(* Logix 5000 project; controller MV vendor 1 type 14 code 217 rev 31.11; software revision 31.00; part 50 of 53 *)
(* tags used below, declared in another part *)
   CC_CIP_BeerMain_Active : DINT;
   CheckTimeMask : INT;
   Delphi_Does_Eng_Func : BOOL;
   enable_comms_to_fv_plc : BOOL;
   MV_BM01_AV01_CIP : BOOL;
   mv_comms_from_cc_plc : MESSAGE;
   mv_comms_from_cc_timer : TIMER;
   MV_COMMS_FROM_FV_PLC : MESSAGE;
   mv_comms_from_mv_routing_plc : MESSAGE;
   mv_comms_to_fv_plc : MESSAGE;
   mv_comms_to_fv_plc_timer : TIMER;
   mv_comms_to_mv_routing_plc : MESSAGE;
   mv_comms_to_mv_routing_plc_timer : TIMER;
   MV_data_file_value_to_move : DINT;
   MV_MV10R : PlantItem;   // MV10R
   MV_MV11R : PlantItem;   // MV11R
   MV_MV12R : PlantItem;   // MV12R
   MV_MV13R : PlantItem;   // MV13R
   MV_MV14R : PlantItem;   // MV14R
   MV_MV15R : PlantItem;   // MV15R
   MV_MV16R : PlantItem;   // MV16R
   MV_MV17R : PlantItem;   // MV17R
   MV_MV18R : PlantItem;   // MV18R
   MV_MV19R : PlantItem;   // MV19R
   MV_MV20_TP_KBEmptying : BOOL;
   MV_MV20R : PlantItem;   // MV20R
   MV_MV21_TP_KBEmptying : BOOL;
   MV_MV21R : PlantItem;   // MV21R
   MV_MV22_TP_KBEmptying : BOOL;
   MV_MV22R : PlantItem;   // MV22R
   MV_MV23R : PlantItem;   // MV23R
   MV_MV30R : PlantItem;   // MV30R
   MV_MV31R : PlantItem;   // MV31R
   MV_MV32R : PlantItem;   // MV32R
   MV_MV33R : PlantItem;   // MV33R
   MV_MV34R : PlantItem;   // MV34R
   MV_MV35R : PlantItem;   // MV35R
   MV_MV7R : PlantItem;   // MV7R
   MV_MV8R : PlantItem;   // MV8R
   MV_MV9R : PlantItem;   // MV9R
   MV_N13 : INT[255];   // PLC>ME Inter PLC comms traf fic inbound
   MV_N14 : INT[255];   // ME>PLC Inter PLC comms traf fic outbound
   MV_N140 : INT[50];   // MV 36, CURRENT FV DATA
   MV_N141 : INT[50];   // MV 37, CURRENT FV DATA
   MV_N142 : INT[50];   // MV 38, CURRENT FV DATA
   MV_N143 : INT[50];   // MV 39, CURRENT FV DATA
   MV_N144 : INT[50];   // MV 40, CURRENT FV DATA
   MV_N145 : INT[50];   // MV 41, CURRENT FV DATA
   MV_N146 : INT[50];   // MV 42, CURRENT FV DATA
   MV_N147 : INT[50];   // MV 43, CURRENT FV DATA
   MV_N148 : INT[50];   // MV 44, CURRENT FV DATA
   MV_N149 : INT[50];   // MV 45, CURRENT FV DATA
   MV_N15 : INT[255];   // COMMS_CTRL Inter PLC comms inte rnal working regs
   MV_N150 : INT[50];   // MV 36, CURRENT FV DATA
   MV_N151 : INT[50];   // MV 47, CURRENT FV DATA
   MV_N15_63_0_OutputBit : BOOL;
   MV_N190 : INT[255];   // Original N File From SLC, No Description Available
   MV_N255 : DINT[255];   // Old Format Checkwords To Keep Delphi Indicating Status Correctly.
   MV_T16 : TIMER[10];
   MV_T191 : TIMER[20];
   MV_T4 : TIMER[20];
   TempChecktime : DINT;
(* MV_Common, continued *)

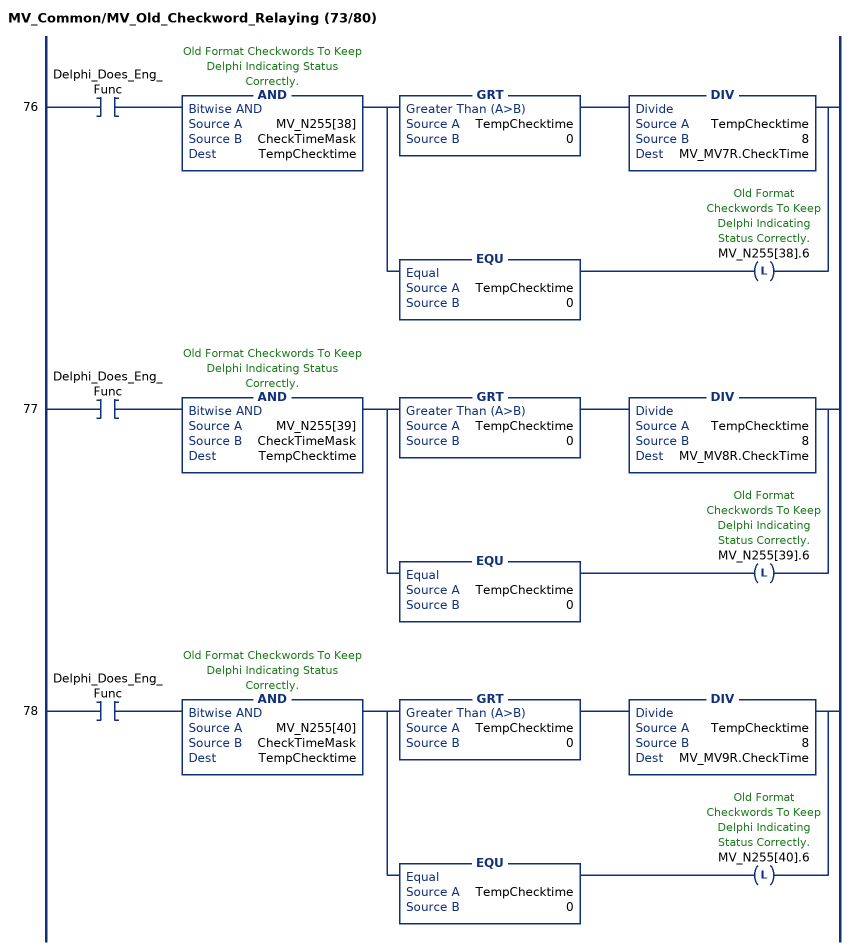
   [picture p1231: MV_Common/MV_Old_Checkword_Relaying rungs 76-78]
   76: XIC(Delphi_Does_Eng_Func)AND(MV_N255[38],CheckTimeMask,TempChecktime)[GRT(TempChecktime,0) DIV(TempChecktime,8,MV_MV7R.CheckTime) ,EQU(TempChecktime,0) OTL(MV_N255[38].6) ];
   77: XIC(Delphi_Does_Eng_Func)AND(MV_N255[39],CheckTimeMask,TempChecktime)[GRT(TempChecktime,0) DIV(TempChecktime,8,MV_MV8R.CheckTime) ,EQU(TempChecktime,0) OTL(MV_N255[39].6) ];
   78: XIC(Delphi_Does_Eng_Func)AND(MV_N255[40],CheckTimeMask,TempChecktime)[GRT(TempChecktime,0) DIV(TempChecktime,8,MV_MV9R.CheckTime) ,EQU(TempChecktime,0) OTL(MV_N255[40].6) ];
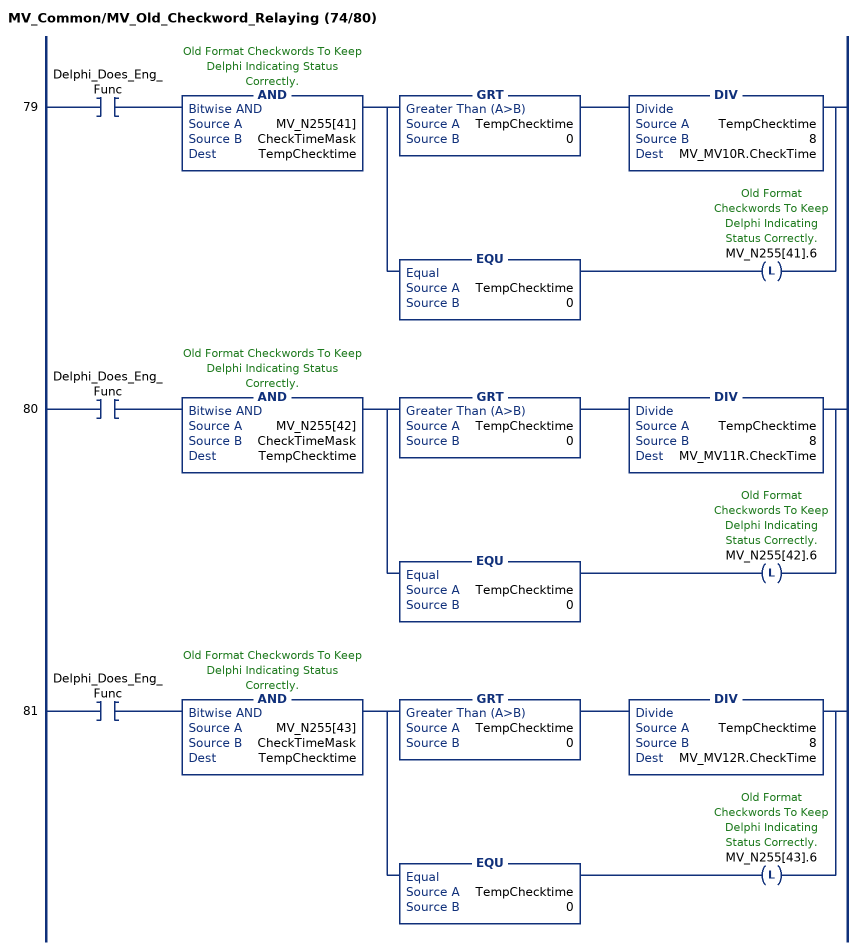
   79: XIC(Delphi_Does_Eng_Func)AND(MV_N255[41],CheckTimeMask,TempChecktime)[GRT(TempChecktime,0) DIV(TempChecktime,8,MV_MV10R.CheckTime) ,EQU(TempChecktime,0) OTL(MV_N255[41].6) ];
   80: XIC(Delphi_Does_Eng_Func)AND(MV_N255[42],CheckTimeMask,TempChecktime)[GRT(TempChecktime,0) DIV(TempChecktime,8,MV_MV11R.CheckTime) ,EQU(TempChecktime,0) OTL(MV_N255[42].6) ];
   81: XIC(Delphi_Does_Eng_Func)AND(MV_N255[43],CheckTimeMask,TempChecktime)[GRT(TempChecktime,0) DIV(TempChecktime,8,MV_MV12R.CheckTime) ,EQU(TempChecktime,0) OTL(MV_N255[43].6) ];
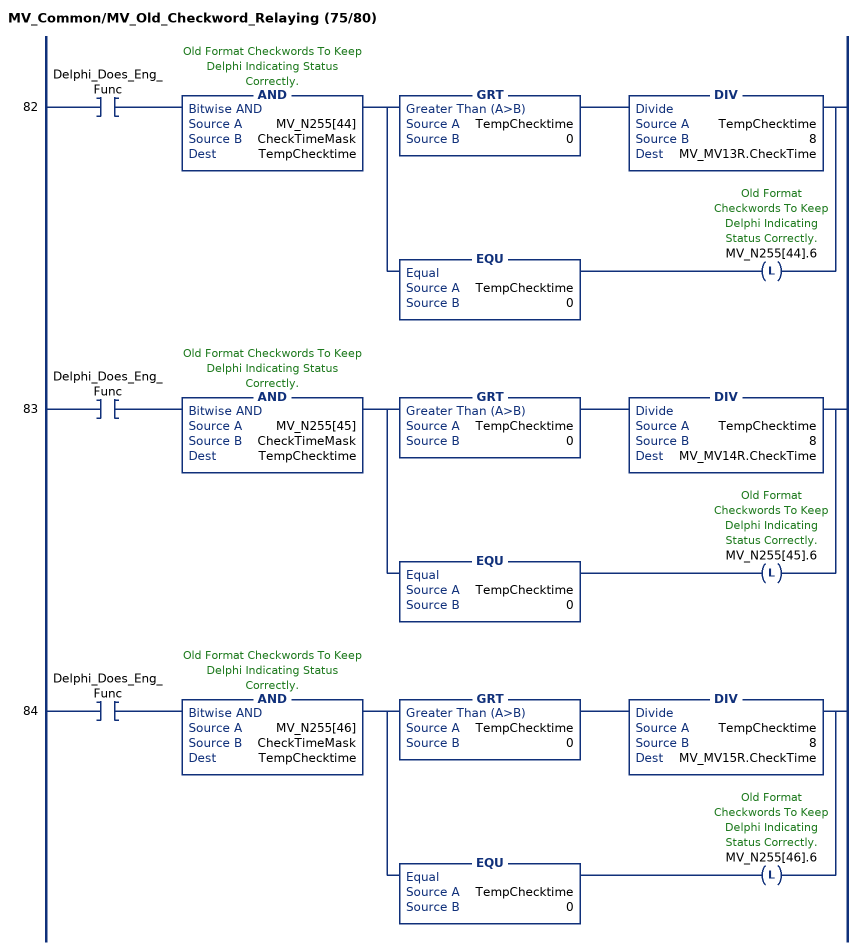
   82: XIC(Delphi_Does_Eng_Func)AND(MV_N255[44],CheckTimeMask,TempChecktime)[GRT(TempChecktime,0) DIV(TempChecktime,8,MV_MV13R.CheckTime) ,EQU(TempChecktime,0) OTL(MV_N255[44].6) ];
   83: XIC(Delphi_Does_Eng_Func)AND(MV_N255[45],CheckTimeMask,TempChecktime)[GRT(TempChecktime,0) DIV(TempChecktime,8,MV_MV14R.CheckTime) ,EQU(TempChecktime,0) OTL(MV_N255[45].6) ];
   84: XIC(Delphi_Does_Eng_Func)AND(MV_N255[46],CheckTimeMask,TempChecktime)[GRT(TempChecktime,0) DIV(TempChecktime,8,MV_MV15R.CheckTime) ,EQU(TempChecktime,0) OTL(MV_N255[46].6) ];
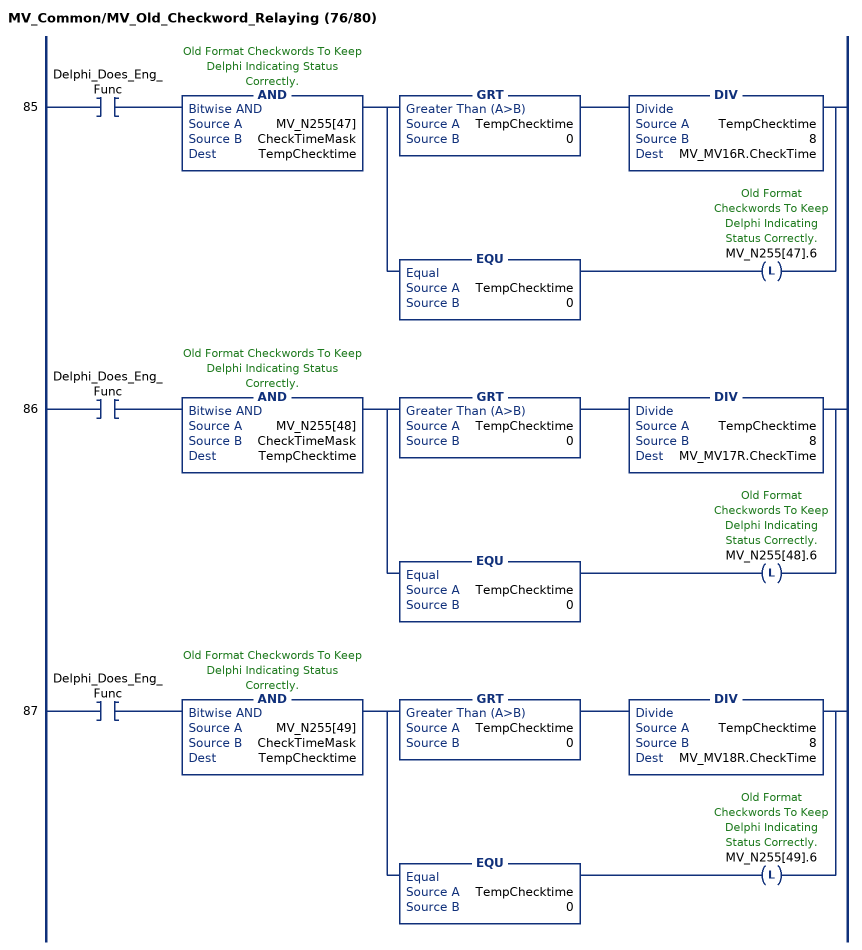
   85: XIC(Delphi_Does_Eng_Func)AND(MV_N255[47],CheckTimeMask,TempChecktime)[GRT(TempChecktime,0) DIV(TempChecktime,8,MV_MV16R.CheckTime) ,EQU(TempChecktime,0) OTL(MV_N255[47].6) ];
   86: XIC(Delphi_Does_Eng_Func)AND(MV_N255[48],CheckTimeMask,TempChecktime)[GRT(TempChecktime,0) DIV(TempChecktime,8,MV_MV17R.CheckTime) ,EQU(TempChecktime,0) OTL(MV_N255[48].6) ];
   87: XIC(Delphi_Does_Eng_Func)AND(MV_N255[49],CheckTimeMask,TempChecktime)[GRT(TempChecktime,0) DIV(TempChecktime,8,MV_MV18R.CheckTime) ,EQU(TempChecktime,0) OTL(MV_N255[49].6) ];
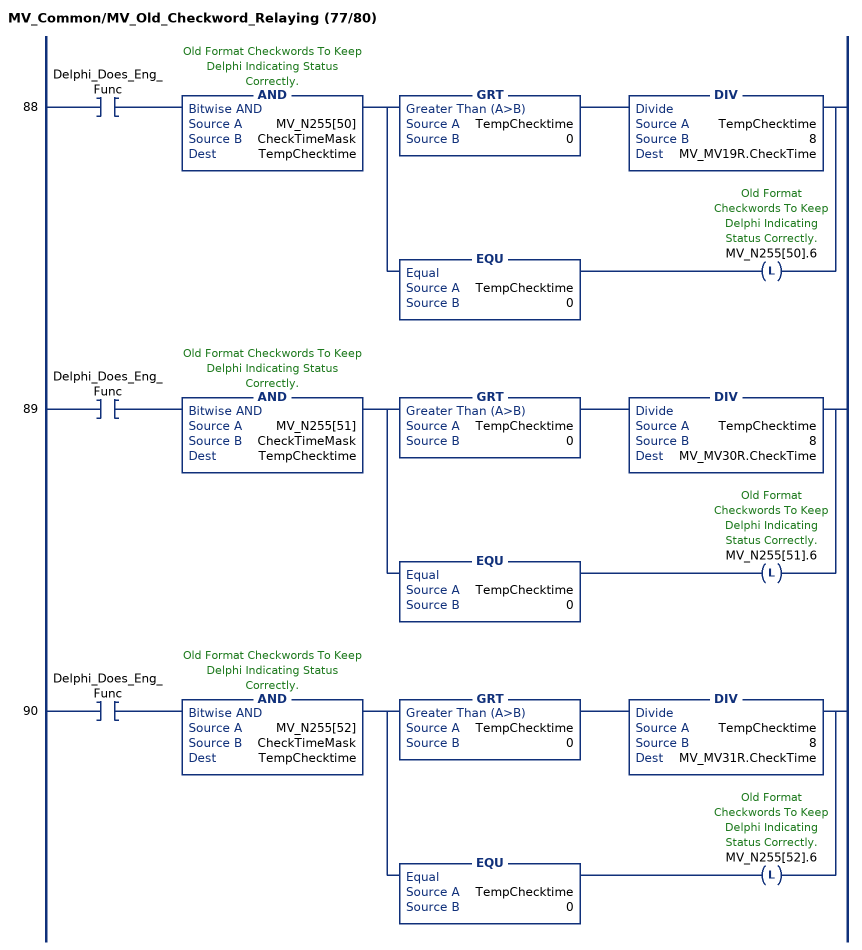
   88: XIC(Delphi_Does_Eng_Func)AND(MV_N255[50],CheckTimeMask,TempChecktime)[GRT(TempChecktime,0) DIV(TempChecktime,8,MV_MV19R.CheckTime) ,EQU(TempChecktime,0) OTL(MV_N255[50].6) ];
   89: XIC(Delphi_Does_Eng_Func)AND(MV_N255[51],CheckTimeMask,TempChecktime)[GRT(TempChecktime,0) DIV(TempChecktime,8,MV_MV30R.CheckTime) ,EQU(TempChecktime,0) OTL(MV_N255[51].6) ];
   90: XIC(Delphi_Does_Eng_Func)AND(MV_N255[52],CheckTimeMask,TempChecktime)[GRT(TempChecktime,0) DIV(TempChecktime,8,MV_MV31R.CheckTime) ,EQU(TempChecktime,0) OTL(MV_N255[52].6) ];
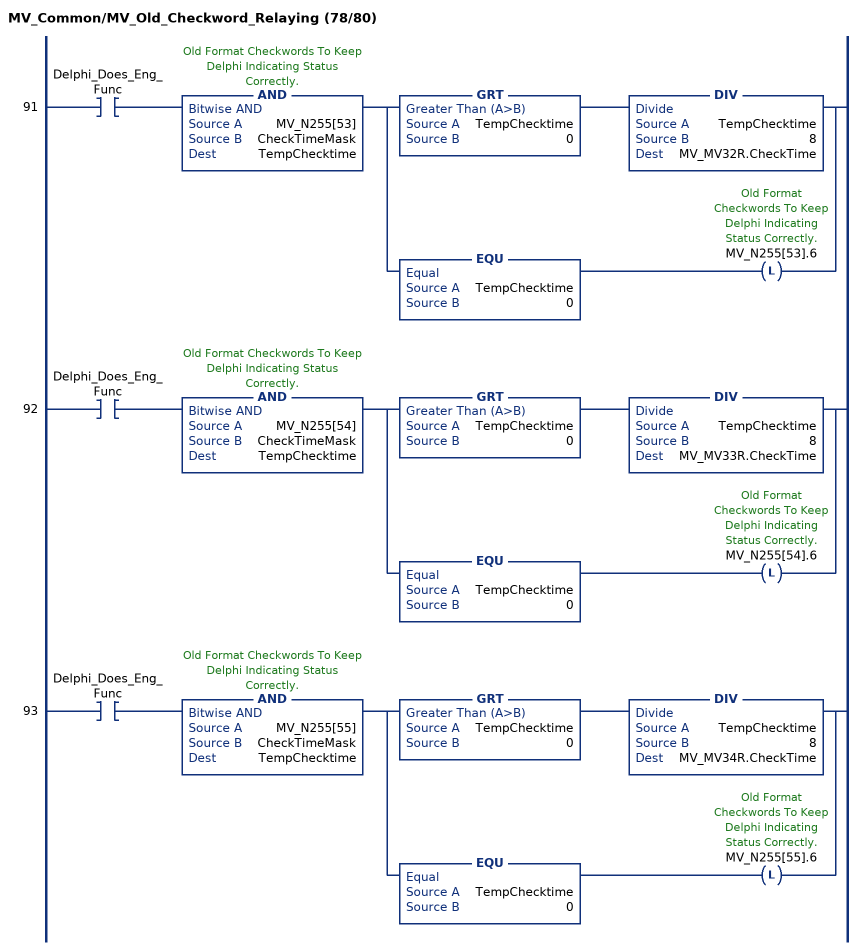
   91: XIC(Delphi_Does_Eng_Func)AND(MV_N255[53],CheckTimeMask,TempChecktime)[GRT(TempChecktime,0) DIV(TempChecktime,8,MV_MV32R.CheckTime) ,EQU(TempChecktime,0) OTL(MV_N255[53].6) ];
   92: XIC(Delphi_Does_Eng_Func)AND(MV_N255[54],CheckTimeMask,TempChecktime)[GRT(TempChecktime,0) DIV(TempChecktime,8,MV_MV33R.CheckTime) ,EQU(TempChecktime,0) OTL(MV_N255[54].6) ];
   93: XIC(Delphi_Does_Eng_Func)AND(MV_N255[55],CheckTimeMask,TempChecktime)[GRT(TempChecktime,0) DIV(TempChecktime,8,MV_MV34R.CheckTime) ,EQU(TempChecktime,0) OTL(MV_N255[55].6) ];
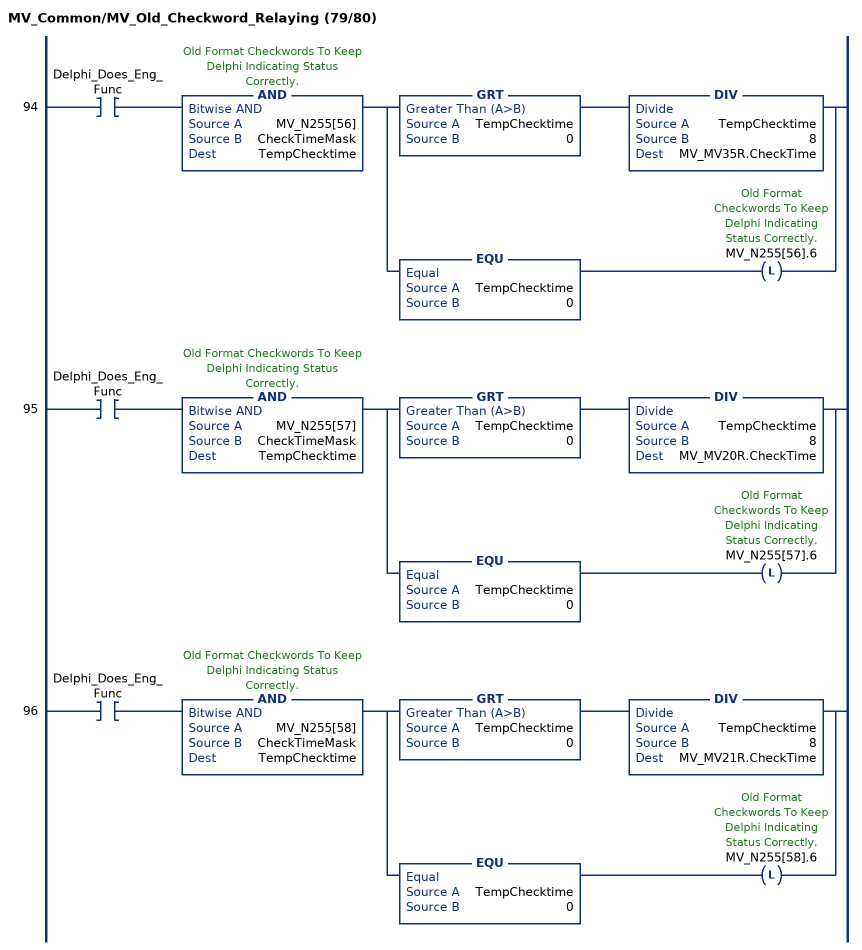
   94: XIC(Delphi_Does_Eng_Func)AND(MV_N255[56],CheckTimeMask,TempChecktime)[GRT(TempChecktime,0) DIV(TempChecktime,8,MV_MV35R.CheckTime) ,EQU(TempChecktime,0) OTL(MV_N255[56].6) ];
   95: XIC(Delphi_Does_Eng_Func)AND(MV_N255[57],CheckTimeMask,TempChecktime)[GRT(TempChecktime,0) DIV(TempChecktime,8,MV_MV20R.CheckTime) ,EQU(TempChecktime,0) OTL(MV_N255[57].6) ];
   96: XIC(Delphi_Does_Eng_Func)AND(MV_N255[58],CheckTimeMask,TempChecktime)[GRT(TempChecktime,0) DIV(TempChecktime,8,MV_MV21R.CheckTime) ,EQU(TempChecktime,0) OTL(MV_N255[58].6) ];
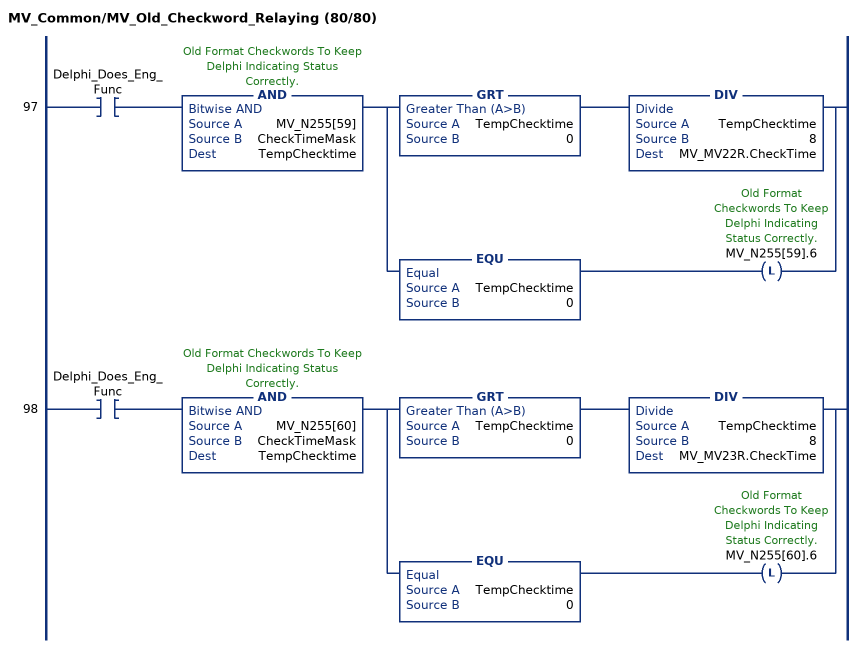
   97: XIC(Delphi_Does_Eng_Func)AND(MV_N255[59],CheckTimeMask,TempChecktime)[GRT(TempChecktime,0) DIV(TempChecktime,8,MV_MV22R.CheckTime) ,EQU(TempChecktime,0) OTL(MV_N255[59].6) ];
   98: XIC(Delphi_Does_Eng_Func)AND(MV_N255[60],CheckTimeMask,TempChecktime)[GRT(TempChecktime,0) DIV(TempChecktime,8,MV_MV23R.CheckTime) ,EQU(TempChecktime,0) OTL(MV_N255[60].6) ];
END_ROUTINE

ROUTINE MV_PLC_COMMS_7   (* ladder *)
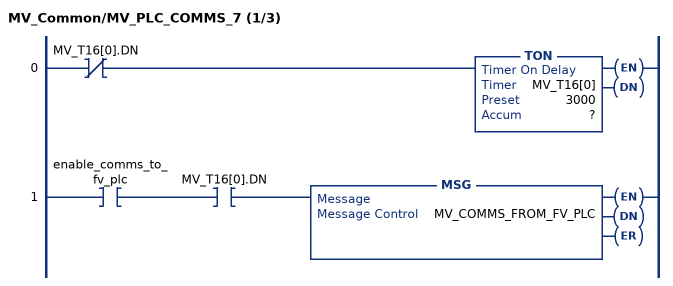
   0: XIO(MV_T16[0].DN)TON(MV_T16[0],?,?);
   1: XIC(enable_comms_to_fv_plc)XIC(MV_T16[0].DN)MSG(MV_COMMS_FROM_FV_PLC);
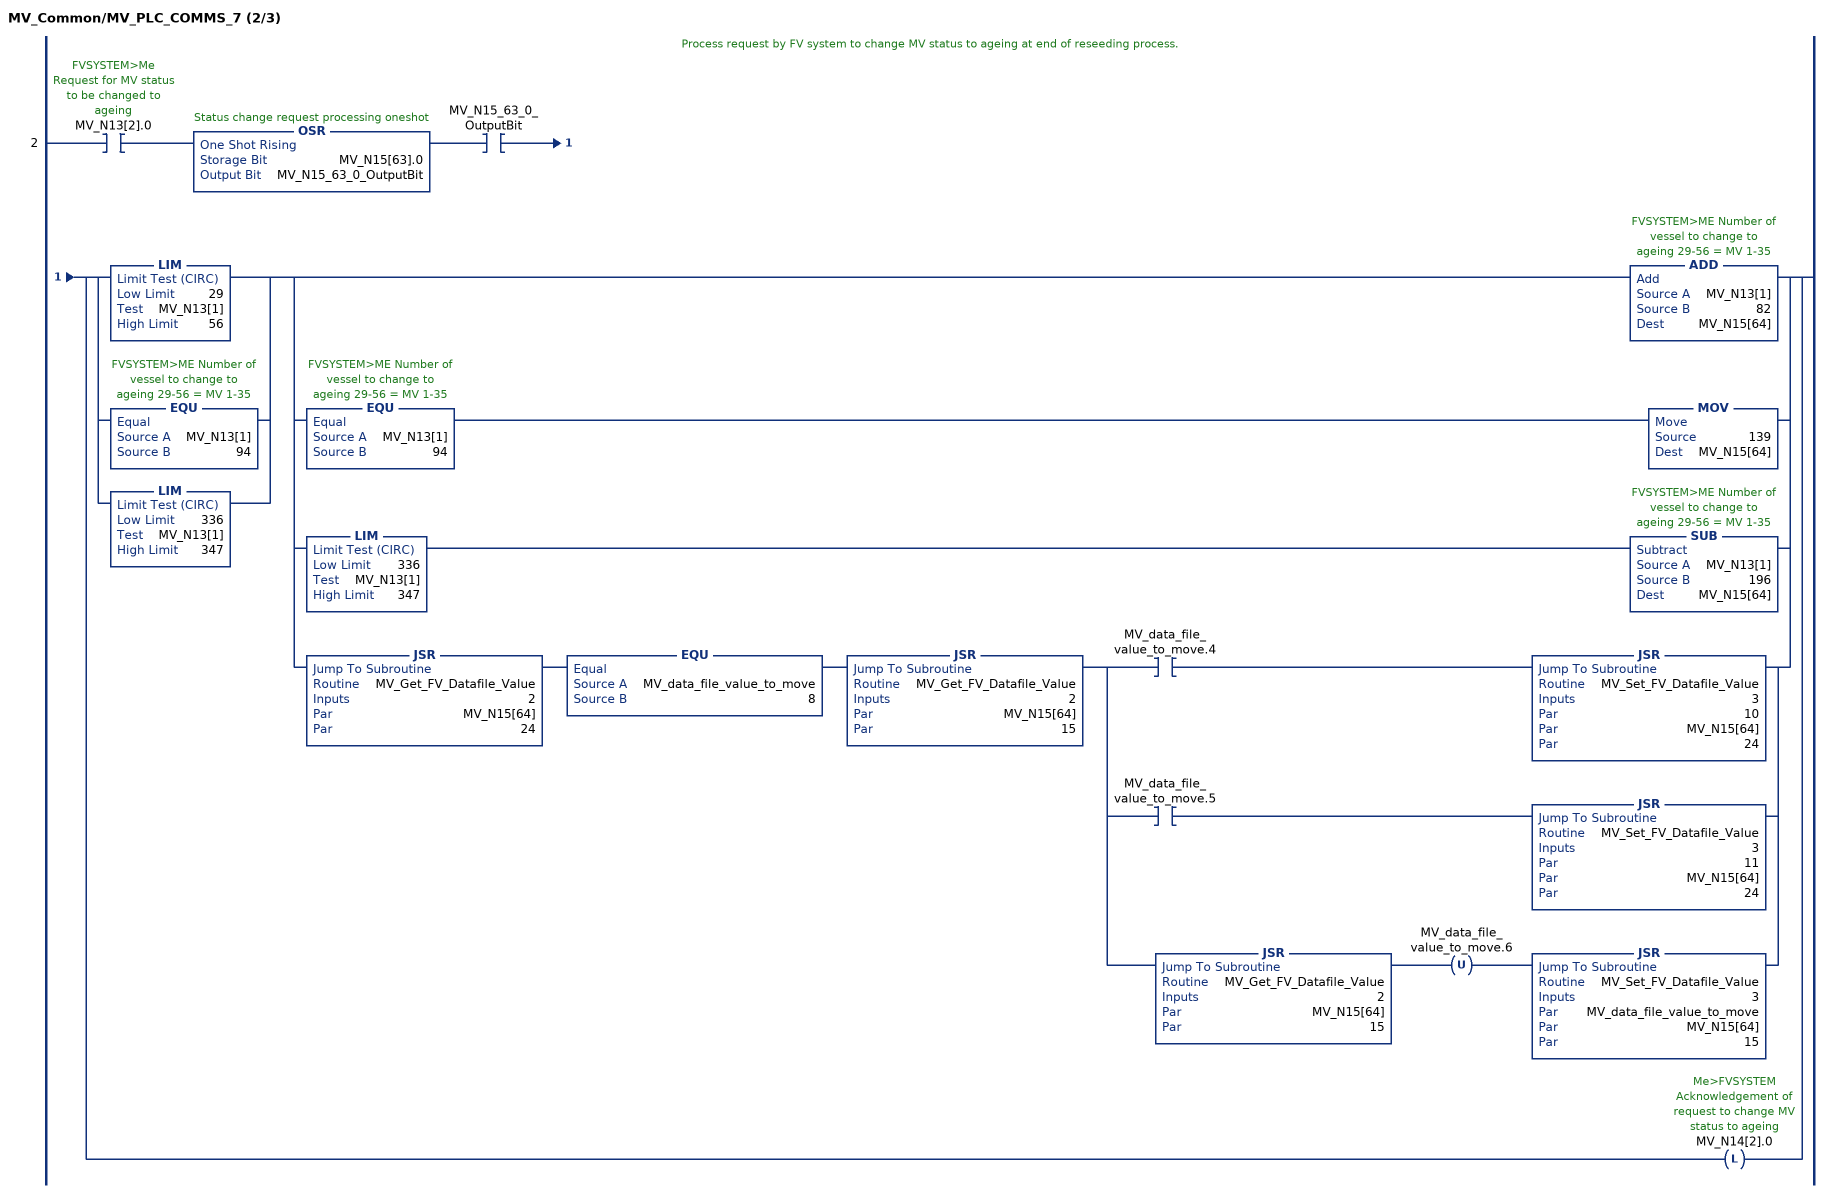
   // Process request by FV system to change MV status to ageing at end of reseeding process.
   2: XIC(MV_N13[2].0)OSR(MV_N15[63].0,MV_N15_63_0_OutputBit)XIC(MV_N15_63_0_OutputBit)[[LIM(29,MV_N13[1],56) ,EQU(MV_N13[1],94) ,LIM(336,MV_N13[1],347) ] [ADD(MV_N13[1],82,MV_N15[64]) ,EQU(MV_N13[1],94) MOV(139,MV_N15[64]) ,LIM(336,MV_N13[1],347) SUB(MV_N13[1],196,MV_N15[64]) ,JSR(MV_Get_FV_Datafile_Value,2,MV_N15[64],24) EQU(MV_data_file_value_to_move,8) JSR(MV_Get_FV_Datafile_Value,2,MV_N15[64],15) [XIC(MV_data_file_value_to_move.4) JSR(MV_Set_FV_Datafile_Value,3,10,MV_N15[64],24) ,XIC(MV_data_file_value_to_move.5) JSR(MV_Set_FV_Datafile_Value,3,11,MV_N15[64],24) ,JSR(MV_Get_FV_Datafile_Value,2,MV_N15[64],15) OTU(MV_data_file_value_to_move.6) JSR(MV_Set_FV_Datafile_Value,3,MV_data_file_value_to_move,MV_N15[64],15) ] ] ,OTL(MV_N14[2].0) ];
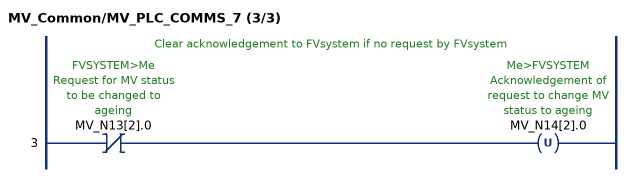
   // Clear acknowledgement to FVsystem if no request by FVsystem
   3: XIO(MV_N13[2].0)OTU(MV_N14[2].0);
END_ROUTINE

ROUTINE MV_PLC_COMMS_9   (* ladder *)
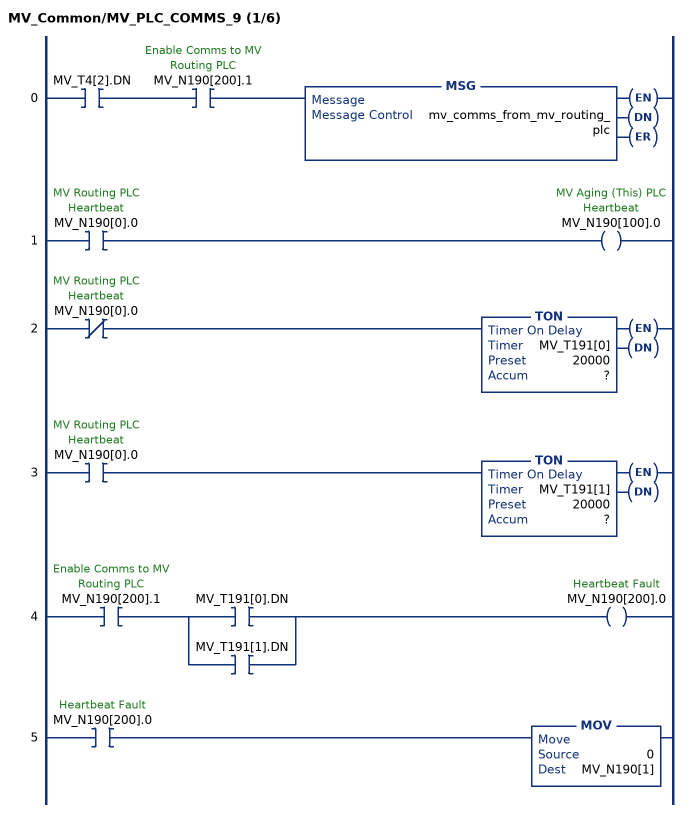
   0: XIC(MV_T4[2].DN)XIC(MV_N190[200].1)MSG(mv_comms_from_mv_routing_plc);
   1: XIC(MV_N190[0].0)OTE(MV_N190[100].0);
   2: XIO(MV_N190[0].0)TON(MV_T191[0],?,?);
   3: XIC(MV_N190[0].0)TON(MV_T191[1],?,?);
   4: XIC(MV_N190[200].1)[XIC(MV_T191[0].DN) ,XIC(MV_T191[1].DN) ]OTE(MV_N190[200].0);
   5: XIC(MV_N190[200].0)MOV(0,MV_N190[1]);
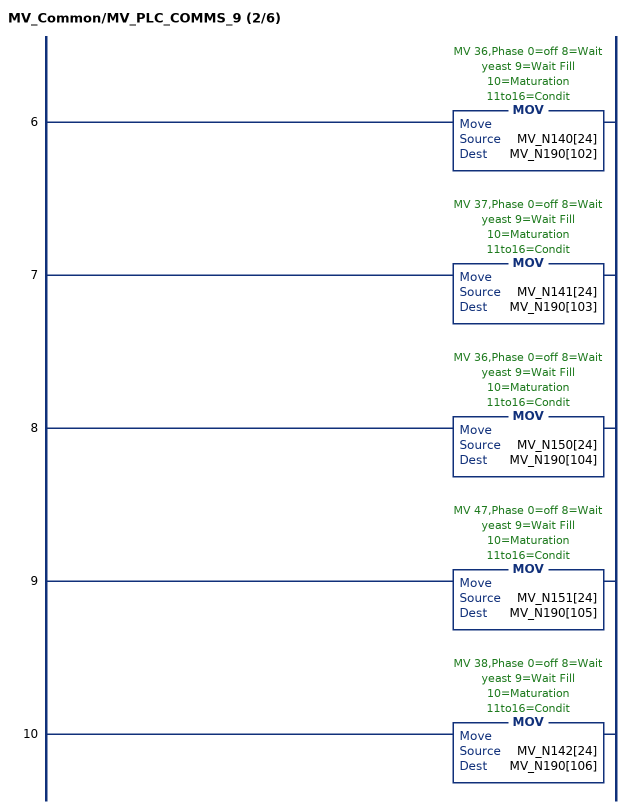
   6: MOV(MV_N140[24],MV_N190[102]);
   7: MOV(MV_N141[24],MV_N190[103]);
   8: MOV(MV_N150[24],MV_N190[104]);
   9: MOV(MV_N151[24],MV_N190[105]);
   10: MOV(MV_N142[24],MV_N190[106]);
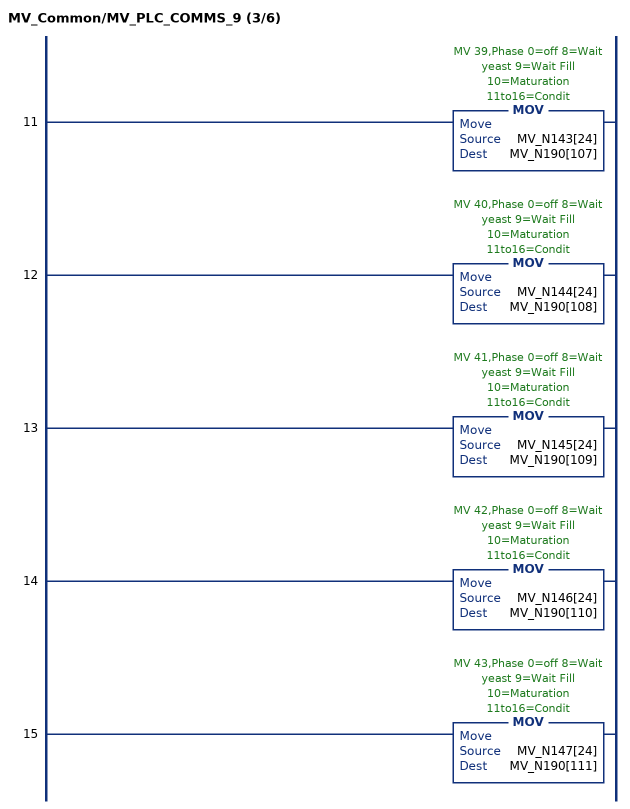
   11: MOV(MV_N143[24],MV_N190[107]);
   12: MOV(MV_N144[24],MV_N190[108]);
   13: MOV(MV_N145[24],MV_N190[109]);
   14: MOV(MV_N146[24],MV_N190[110]);
   15: MOV(MV_N147[24],MV_N190[111]);
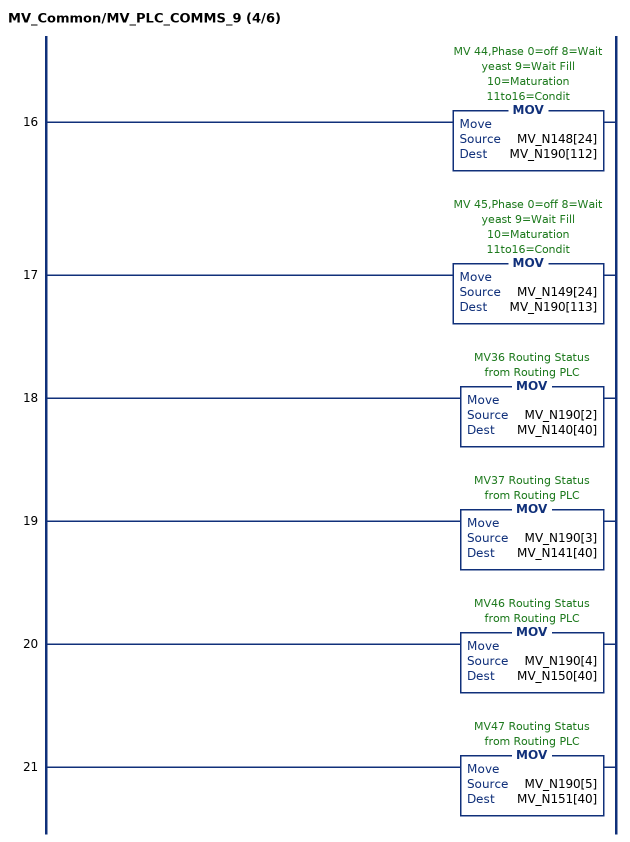
   16: MOV(MV_N148[24],MV_N190[112]);
   17: MOV(MV_N149[24],MV_N190[113]);
   18: MOV(MV_N190[2],MV_N140[40]);
   19: MOV(MV_N190[3],MV_N141[40]);
   20: MOV(MV_N190[4],MV_N150[40]);
   21: MOV(MV_N190[5],MV_N151[40]);
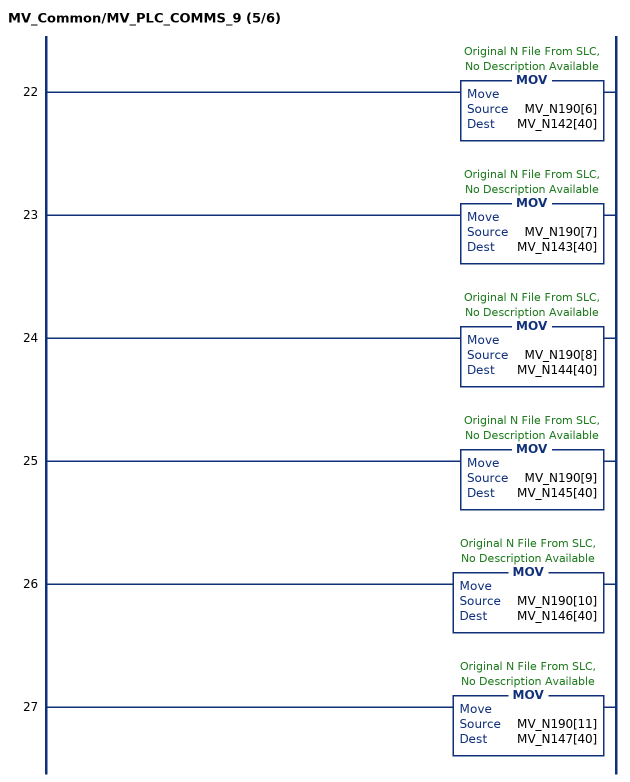
   22: MOV(MV_N190[6],MV_N142[40]);
   23: MOV(MV_N190[7],MV_N143[40]);
   24: MOV(MV_N190[8],MV_N144[40]);
   25: MOV(MV_N190[9],MV_N145[40]);
   26: MOV(MV_N190[10],MV_N146[40]);
   27: MOV(MV_N190[11],MV_N147[40]);
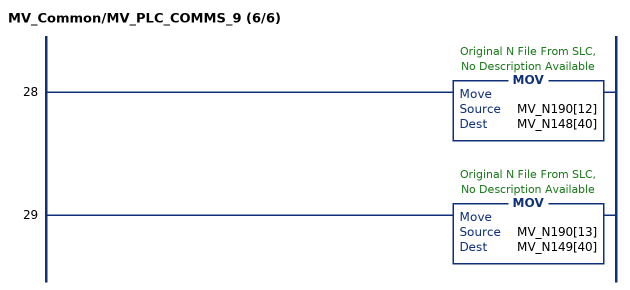
   28: MOV(MV_N190[12],MV_N148[40]);
   29: MOV(MV_N190[13],MV_N149[40]);
END_ROUTINE

ROUTINE MV_PLC_COMMS_Write_Replacements   (* ladder *)
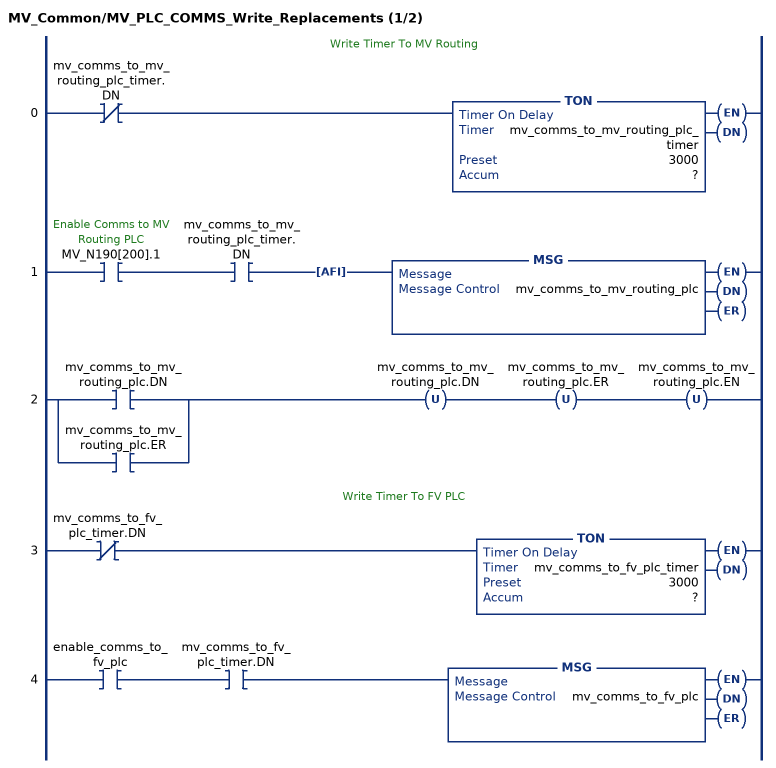
   // Write Timer To MV Routing
   0: XIO(mv_comms_to_mv_routing_plc_timer.DN)TON(mv_comms_to_mv_routing_plc_timer,?,?);
   1: XIC(MV_N190[200].1)XIC(mv_comms_to_mv_routing_plc_timer.DN)AFI()MSG(mv_comms_to_mv_routing_plc);
   2: [XIC(mv_comms_to_mv_routing_plc.DN) ,XIC(mv_comms_to_mv_routing_plc.ER) ]OTU(mv_comms_to_mv_routing_plc.DN)OTU(mv_comms_to_mv_routing_plc.ER)OTU(mv_comms_to_mv_routing_plc.EN);
   // Write Timer To FV PLC
   3: XIO(mv_comms_to_fv_plc_timer.DN)TON(mv_comms_to_fv_plc_timer,?,?);
   4: XIC(enable_comms_to_fv_plc)XIC(mv_comms_to_fv_plc_timer.DN)MSG(mv_comms_to_fv_plc);
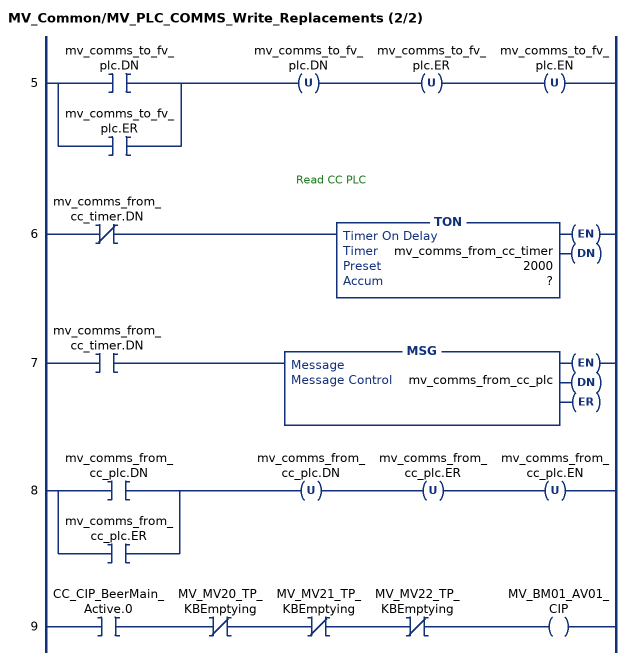
   5: [XIC(mv_comms_to_fv_plc.DN) ,XIC(mv_comms_to_fv_plc.ER) ]OTU(mv_comms_to_fv_plc.DN)OTU(mv_comms_to_fv_plc.ER)OTU(mv_comms_to_fv_plc.EN);
   // Read CC PLC
   6: XIO(mv_comms_from_cc_timer.DN)TON(mv_comms_from_cc_timer,?,?);
   7: XIC(mv_comms_from_cc_timer.DN)MSG(mv_comms_from_cc_plc);
   8: [XIC(mv_comms_from_cc_plc.DN) ,XIC(mv_comms_from_cc_plc.ER) ]OTU(mv_comms_from_cc_plc.DN)OTU(mv_comms_from_cc_plc.ER)OTU(mv_comms_from_cc_plc.EN);
   9: XIC(CC_CIP_BeerMain_Active.0)XIO(MV_MV20_TP_KBEmptying)XIO(MV_MV21_TP_KBEmptying)XIO(MV_MV22_TP_KBEmptying)OTE(MV_BM01_AV01_CIP);
END_ROUTINE
